(* CODESYS project CanOpen.project
   Title: Opus30
   Version: 1.0.0.0
   Author: Marcus Adolfi
   Company: Schneider Electric

Project tree, tasks and I/O mapping:
  MyController : TM241CE40T/U, Schneider Electric, order no. TM241CE40T/U, version 4.0.2.20
    application Application
      libraries: SysTime, 3.4.1.20 (System)
      task MAST (cyclic, interval 10 ms, priority 15, watchdog 100 ms x 1) calls R00_main
      task VISU_TASK (cyclic, interval 100 ms, priority 30) calls VisuElems.Visu_Prg
      task Task1ms (cyclic, interval 1 ms, priority 1) calls F04_foto, D04_foto, S06_seguranca
      global variables GVL
      01_Machine/
        program R06_principal [LD]
        program R01_firstScan [LD]
        program R05_comando [LD]
        program R21_estatistica [ST]
        program R22_velocMedia [ST]
        program R98_paramFab [ST]
        program R20_acessorios [LD]
        program R99_calcTempos [ST]
        program R00_main [LD]
      Structs/
        data type _exec_bits
        data type _eixo_drive
        data type _eixo_home
        data type _eixo_auto
        data type _receita
        data type _eixo
        data type _bio
        data type _oee
        data type _prev
      05_IHM/
        program I02_alarmes [ST]
        program I07_procedimento [LD]
        program I06_textoConfirma [LD]
        program I01_geral [LD]
        program I03_mensagens [ST]
      02_Filme/
        program F99_calculo [ST]
        program F03_auto [LD]
        program F01_geral [LD]
        program F04_foto [LD]
      global variables PersistentVars
      03_Selagem/
        program S02_home [LD]
        program S99_calculo [ST]
        program S06_seguranca [LD]
        program S01_geral [LD]
        program S03_auto [LD]
      global variables IHM
      Symbol configuration
      04_Disco/
        program D99_calculo [ST]
        program D03_auto [LD]
        program D04_foto [LD]
      function HiddenPOU [ST]
      Visu/
        visualisation Info
        visualisation Main
      10_Relogio/
        function block GetDateAndTime [CFC]
        function block SetDateAndTime [CFC]
        program AjustaDataHora [LD]
      image pool Imagens
      11_FB/
        function block RTO [ST]
      06_bio/
        program B01_controle [ST]
        program B02_data [ST]
      07_dados/
        program D01_data [ST]
        program D02_clean [ST]
        program D03_view [ST]
        program D04_controleView [ST]
      08_manut/
        program U01_controle [ST]
        program U02_soma [ST]
        program U03_reset [ST]
        program U04_view [ST]
        program U00_valoresMax [ST]
    Cartridge_1 : Cartridge, Schneider Electric, version 4.0.2.20
    Cartridge_2 : Cartridge, Schneider Electric, version 4.0.2.20
    IO_Bus : IO bus - TM3, Schneider Electric, version 4.0.2.20
    COM_Bus : COM bus, Schneider Electric, version 4.0.2.20
    Ethernet_1 : Ethernet Network, Schneider Electric, version 4.0.2.20
        settings: IPAddress = [192, 168, 1, 10]; SubnetMask = [255, 255, 255, 0]; WebServer = TRUE; FTP Server = TRUE; SoMachine Protocol = TRUE; Modbus Server = TRUE; NetManage Protocol = TRUE; SNMP protocol = TRUE; WebVisu protocol = TRUE
    Serial_Line_1 : Serial line, Schneider Electric, version 4.0.2.20
      SoMachine_Network_Manager : SoMachine-Network Manager, Schneider Electric, version 4.0.0.2
    Serial_Line_2 : Serial line, Schneider Electric, version 4.0.2.20
      Modbus_Manager : Modbus Manager, Schneider Electric, version 4.0.0.7
    DI : Digital Inputs, Schneider Electric, version 4.0.2.20
        input  i_fotoFilme : BOOL  // IDW0.I0
        input  i_selagFechado : BOOL  // IDW0.I1
        input  i_fotoDisco : BOOL  // IDW0.I2
        input  i_segProduto : BOOL  // IDW0.I3
        input  i_fechamDisco : BOOL  // IDW0.I4
        input  i_selagAberto : BOOL  // IDW0.I5
        input  i_paradaCorte : BOOL  // IDW0.I6
        input  i_relePortaSeg : BOOL  // IDW0.I7
        input  i_segParada : BOOL  // IDW0.I8
        input  i_btReset : BOOL  // IDW0.I9
        input  i_releEmergencia : BOOL  // IDW0.I10
        input  i_marchaAutomatica : BOOL  // IDW0.I11
        input  i_botaoCiclo : BOOL  // IDW0.I12
        input  i_falhaTemperatura : BOOL  // IDW0.I13
        input  i_falhaImpressora : BOOL  // IDW0.I14
        unmapped channels: IDW0, IB1
    DQ : Digital Outputs, Schneider Electric, version 4.0.2.20
        output o_corte : BOOL  // QW0.Q6
        output o_impressao : BOOL  // QW0.Q7
        output o_compressor : BOOL  // QW0.Q9
        output o_injecaoAr : BOOL  // QW0.Q10
        output o_liberaFilme : BOOL  // QW0.Q13
        output qbDQ_QB1 : BYTE  // QB1
        unmapped channels: QW0
    Counters : Counters, Schneider Electric, version 4.0.2.20
    Pulse_Generators : Pulse Generators, Schneider Electric, version 4.0.2.20
        settings: InstanceNumber = 0; Instance name = 'filme_PTO'; Temporary Instance name = 'filme_PTO'; InstanceNumber = 1; Instance name = 'selag_PTO'; Temporary Instance name = 'selag_PTO'
  HMISTU855 : HMIS5T, Schneider Electric, order no. HMIS5T, version 3.5.3.46
    HMI Application
    Ethernet
      SoMachine_Network_Manager2 : SoMachine-Network Manager, Schneider Electric, version 4.0.0.2
    USB
      SoMachine_Network_Manager3 : SoMachine-Network Manager, Schneider Electric, version 4.0.0.2
    COM1
      SoMachine_Network_Manager1 : SoMachine-Network Manager, Schneider Electric, version 4.0.0.2
  6c0f7fb6-600b-4c93-9262-20cdc603757e
  text list GlobalTextList
  5ce3da45-db07-42e7-a21c-a00fff4ed8f6|C:\_Clientes\Opuspac\Doc\Figuras\Botao.png
  5ce3da45-db07-42e7-a21c-a00fff4ed8f6|C:\_Clientes\Opuspac\Doc\Figuras\Botao_ps.png
  5ce3da45-db07-42e7-a21c-a00fff4ed8f6|C:\_Clientes\Opuspac\Doc\Figuras\LogoOpus.jpg
*)

// MyController/Application/Structs/_exec_bits
TYPE _exec_bits :
STRUCT
	RQ					: BOOL;
	IP					: BOOL;
	DN					: BOOL;
	Fase				: DINT;
	Mask				: DINT;
END_STRUCT
END_TYPE

// MyController/Application/Structs/_eixo_drive
TYPE _eixo_drive :
STRUCT
	falha			: MC_ReadAxisError_PTO;
	posicao			: MC_ReadActualPosition_PTO;
	power			: MC_Power_PTO;
	reset			: MC_Reset_PTO;
	status			: MC_ReadMotionState_PTO;
	stop			: MC_Stop_PTO;
END_STRUCT
END_TYPE

// MyController/Application/Structs/_eixo_home
TYPE _eixo_home :
STRUCT
	RQ					: BOOL;
	IP					: BOOL;
	DN					: BOOL;
	Fase				: DINT;
	Mask				: DINT;
	movVeloc			: MC_MoveVelocity_PTO;
	movRelat			: MC_MoveRelative_PTO;
	movStop				: ARRAY[1..2] OF MC_Stop_PTO;
	setPos				: MC_SetPosition_PTO;
END_STRUCT
END_TYPE

// MyController/Application/Structs/_eixo_auto
TYPE _eixo_auto :
STRUCT
	movVeloc					: MC_MoveVelocity_PTO;
	movAbs						: ARRAY[0..2] OF MC_MoveAbsolute_PTO;
	movRelat					: ARRAY[0..2] OF MC_MoveRelative_PTO;
	movStop						: MC_Stop_PTO;
	setPos						: MC_SetPosition_PTO;
END_STRUCT
END_TYPE

// MyController/Application/Structs/_receita
TYPE _receita :
STRUCT
	inicioAtraso				: DINT;

	// Filme
	filmeExtra					: BOOL;
	filmeMmAposFoto				: DINT;
	filmeMmExtra				: DINT;
	
	// Disco
	discoMmAposFoto				: DINT;
	discoAtraso					: DINT;
END_STRUCT
END_TYPE

// MyController/Application/Structs/_eixo
TYPE _eixo :
STRUCT
	auto				: _eixo_auto;
	home				: _eixo_home;
	drive				: _eixo_drive;
	falha				: BOOL;
	posicaoAtual		: DINT;
	calcula				: BOOL;
END_STRUCT
END_TYPE

// MyController/Application/Structs/_bio
TYPE _bio :
STRUCT
	login						: WSTRING:= "";
	loginData					: BOOL;
	bioData						: ARRAY [0..49] OF DINT;
	bioHora						: ARRAY [0..49] OF DINT;
	bioMin						: ARRAY [0..49] OF DINT;
	bioUser						: ARRAY [0..49] OF WSTRING;
	bioGui						: ARRAY [0..49] OF BOOL;
	iz							: DINT:= 0;
END_STRUCT
END_TYPE

// MyController/Application/Structs/_oee
TYPE _oee :
STRUCT
	produtividade				: ARRAY [0..30] OF REAL;
	diaProduzido				: ARRAY [0..30] OF UINT;
	horasProduzidas				: ARRAY [0..30] OF DINT;
	minProduzidos				: ARRAY [0..30] OF DINT;
	diaProduzindo				: DINT;
	mesProduzindo				: DINT;
	anoProduzindo				: DINT;
	backUpdia					: BOOL;
	pontIhm						: ARRAY [0..30] OF BOOL;
	diaProd						: DINT;
END_STRUCT
END_TYPE

// MyController/Application/Structs/_prev
TYPE _prev :
STRUCT
	M_ciclosMax	 				: ARRAY[ 0..7] OF  DINT;
	ciclos						: ARRAY[ 0..7] OF  DINT;
	msg							: ARRAY[ 0..7] OF  BOOL;
	habilita					: ARRAY[ 0..7] OF BOOL;
END_STRUCT
END_TYPE

// MyController/Application/GVL
VAR_GLOBAL
	// transições
	psBtCiclo					: BOOL;

	// Variaveis gerais
	alarmeReset					: BOOL;
	alarmeResetInd				: BOOL;
	alarmeResetBtn				: BOOL;
	alwaysOff					: BOOL;
	alwaysOn					: BOOL;
	arOK						: BOOL;
	biometricoOk				: BOOL;
	calcGeral					: BOOL;
	calcTempos					: BOOL;
	comandoOff					: BOOL;
	contaReset					: BOOL;
	emergOk						: BOOL;
	estatReset					: BOOL;
	existeAlarme				: BOOL;
	falhaImpressora				: BOOL;
	falhaProduto				: BOOL;
	falhaSensorProd				: BOOL;
	falhaTemperatura			: BOOL;
	firstScan					: BOOL;
	injecaoTpoOff				: BOOL;
	liberaCiclo					: BOOL;
	livreComando				: BOOL;
	livreStart					: BOOL;
	modoAutomatico				: BOOL;					
	pisca						: BOOL;
	piscaRapido					: BOOL;
	primeiroCiclo				: BOOL;
	setAmpola					: BOOL;
	tpoDisco					: TIME;
	tpoInicio					: TIME;
	tpoInjecao					: TIME;
	tpoSelagem					: TIME;
	
	
	
	TL_inicializa				: TON;
	TL_disco					: TON;
	TF_corte					: TON;
	
	acopla						: _exec_bits;
	ciclo						: _exec_bits;
	comando						: _exec_bits;
	compressor					: _exec_bits;
	conta						: _exec_bits;
	corte						: _exec_bits;
	injecaoAr					: _exec_bits;
	media						: _exec_bits;
	mudaReceita					: _exec_bits;
	principal					: _exec_bits;
	vidaUtil					: _exec_bits;
	
	// Alimentador de Blisters
	msgPrimeiro					: BOOL;
	limpaDados					: BOOL;
	procedimento				: ARRAY[0..2] OF _exec_bits;

	
	// Variaveis Filme
	filme						: _eixo;
	filmeMove					: ARRAY[0..2] OF _exec_bits;
	filmeParaImed				: BOOL;
	filmeVeloc					: DINT;
	filmeExtra					: BOOL;
	filmeFotoOk					: BOOL;
	filmePulsosAposFoto			: DINT;
	filmePulsosExtra			: DINT;
	filmePulsosMm				: REAL;
	filmePreso					: _exec_bits;
	
	// Variaveis Selagem
	selag						: _eixo;
	selagAbre					: _exec_bits;
	selagFecha					: _exec_bits;
	selagVeloc					: DINT;
	selagVelocHome				: DINT;
	selagPulsosMm				: REAL;
	selagPulsosFechar			: DINT;

	// Variaveis Disco
	disco						: _eixo;
	discoMove					: _exec_bits;
	discoParaImed				: BOOL;
	discoVeloc					: DINT;
	discoPulsosMm				: REAL;
	discoPulsosAposFoto			: DINT;
	
	// Variaveis Visualization
	vsBtStart					: BOOL;
	vsMarchaAutomatica			: BOOL;
	
	
    //Sincroniza e ajusta o relógio da IHM
	AnoSet						: UINT;
	ClkScan						: BOOL;
	AjustaHora					: BOOL;
	MesSet						: UINT;
	DiaSet						: UINT;
	HoraSet						: UINT;
	MinutoSet					: UINT;
	SegundoSet					: UINT;
	AnoAtual					: UINT;
	MesAtual					: UINT;
	DiaAtual					: UINT;
	HoraAtual					: UINT;
	MinutoAtual					: UINT;
	SegundoAtual				: UINT;	
	sink						: BOOL;

	
(*	=================== ALARMES ===================
	Obs: alarme[0]- Não utilizado
*)
	alarme						: ARRAY[0..50] OF BOOL;
	alarmes						: _exec_bits;
	mensagem					: ARRAY[0..50] OF BOOL;
	numAlarme					: SINT;
END_VAR

// MyController/Application/PersistentVars
VAR_GLOBAL PERSISTENT RETAIN
	versaoSoftware				: REAL:= 1.00;
	pi							: REAL:= 3.1415926;
	paramFab					: BOOL:= TRUE;
	contaAtual					: DINT;
	contaGeral					: DINT;
	contaSet					: DINT;
	numReceita					: SINT;
	
	M_tpoInjecaoAr				: DINT:= 99;
	M_produtMedio				: DINT:= 70;
	M_tpoFormato				: TIME:= T#280MS;
	
	// Informações
	infoTpoEnergHrs				: DINT;
	infoTpoEnergMin				: DINT;
	infoTpoProdHrs				: DINT;
	infoTpoProdMin				: DINT;
	
	// Filme
	M_filmePulsosVolta			: DINT:= 1600;
	M_diamRolo					: DINT:= 34;
	M_filmeVeloc				: DINT:= 40;
	M_filmeAcel					: DINT:= 200;
	M_filmeDecel				: DINT:= 100;
	
	// Disco
	M_discoPulsosVolta			: DINT:= 6400;
	M_diamDisco					: DINT:= 166;
	M_discoVeloc				: DINT:= 4;
	M_discoAcel					: DINT:= 150;
	M_discoDecel				: DINT:= 150;
	
	// Selagem
	M_selagPulsosVolta			: DINT:= 20000;
	M_selagVelocHome			: DINT:= 20;
	M_selagVeloc				: DINT:= 100;
	M_selagTpoSelagem			: DINT:= 20;
	M_selagPosFecha				: DINT:= 789;
	M_selagAcel					: DINT:= 40;
	M_selagDecel				: DINT:= 40;
	
	// Receita
	Rc							: ARRAY[0..3] OF _receita;
	Fb							: ARRAY[0..3] OF _receita;
	
	// IHM
	ihm_procedCurto				: BOOL;
	
	// Digital
	digital						: _bio;
	iz							: DINT;
	
	// biometria
	ihm_digitalInstalado		: BOOL;
	
	// Dados
	dados						: _oee;
	indPainel					: DINT:= 0;
	indSub						: BOOL;
	indSoma						: BOOL;
	panData						: ARRAY [0..08] OF DINT;
	panProd						: ARRAY [0..08] OF REAL;
	panHora						: ARRAY [0..08] OF DINT;
	panMin						: ARRAY [0..08] OF DINT;
	pt							: DINT:= 0;
	pa							: DINT;
	
	// Vida Util
	util						: _prev; 
END_VAR

// MyController/Application/IHM
VAR_GLOBAL
	ihm_alarme					: ARRAY[0..50] OF BOOL;
	ihm_alarmeReset				: BOOL;
	ihm_alarmeResetInd			: BOOL;
	ihm_bannerConfirma			: BOOL;
	ihm_bannerMensagem			: BOOL;
	ihm_carregaFabrica			: BOOL;
	ihm_confirmaV				: BOOL;
	ihm_confirmaX				: BOOL;
	ihm_contaAtual				: DINT;
	ihm_contaGeral				: DINT;
	ihm_contaReset				: BOOL;
	ihm_entrada					: ARRAY[0..23] OF BOOL;
	ihm_estatReset				: BOOL;
	ihm_mensagem				: DINT;
	ihm_numReceita				: SINT;
	ihm_preso					: BOOL;
	ihm_produtMedio				: REAL;
	ihm_telaHome				: BOOL;
	ihm_salvaFabrica			: BOOL;
	ihm_saida					: ARRAY[0..15] OF BOOL;
	ihm_selagHome				: BOOL;
	ihm_telaAtual				: INT;
	ihm_textoConfirma			: DINT;
	ihm_textoProced				: DINT;
	ihm_velocMedida				: DINT;
	ihm_visibPhone				: BOOL;
	ihm_setUpAmpola				: BOOL;
	
	// Produtividade
	ihm_backUpProdutividade		: BOOL;
	
	
	ihm_digitalHabilitado		: BOOL;
	ihm_usuarioLoggado			: BOOL;
	ihm_realizaBackup 			: BOOL;	
	
	// Vida Util 
	ihm_resetCiclos				: ARRAY[0..7] OF BOOL;
END_VAR

// MyController/Application/01_Machine/R00_main
PROGRAM R00_main
VAR
END_VAR

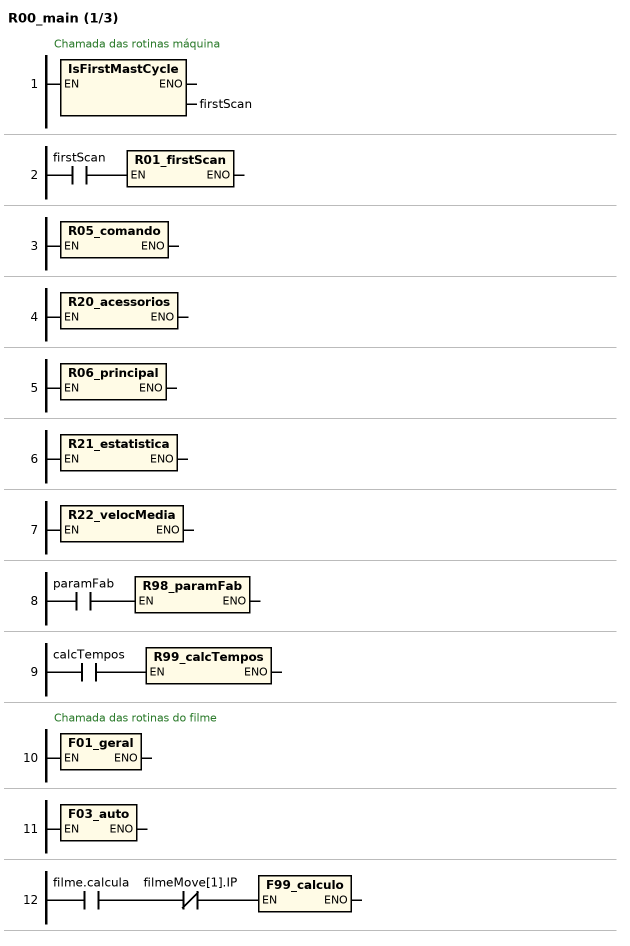
// NETWORK 1
// Chamada das rotinas máquina
firstScan := IsFirstMastCycle();

// NETWORK 2
IF firstScan THEN R01_firstScan(); END_IF

// NETWORK 3
R05_comando();

// NETWORK 4
R20_acessorios();

// NETWORK 5
R06_principal();

// NETWORK 6
R21_estatistica();

// NETWORK 7
R22_velocMedia();

// NETWORK 8
IF paramFab THEN R98_paramFab(); END_IF

// NETWORK 9
IF calcTempos THEN R99_calcTempos(); END_IF

// NETWORK 10
// Chamada das rotinas do filme
F01_geral();

// NETWORK 11
F03_auto();

// NETWORK 12
IF filme.calcula AND NOT filmeMove[1].IP THEN F99_calculo(); END_IF

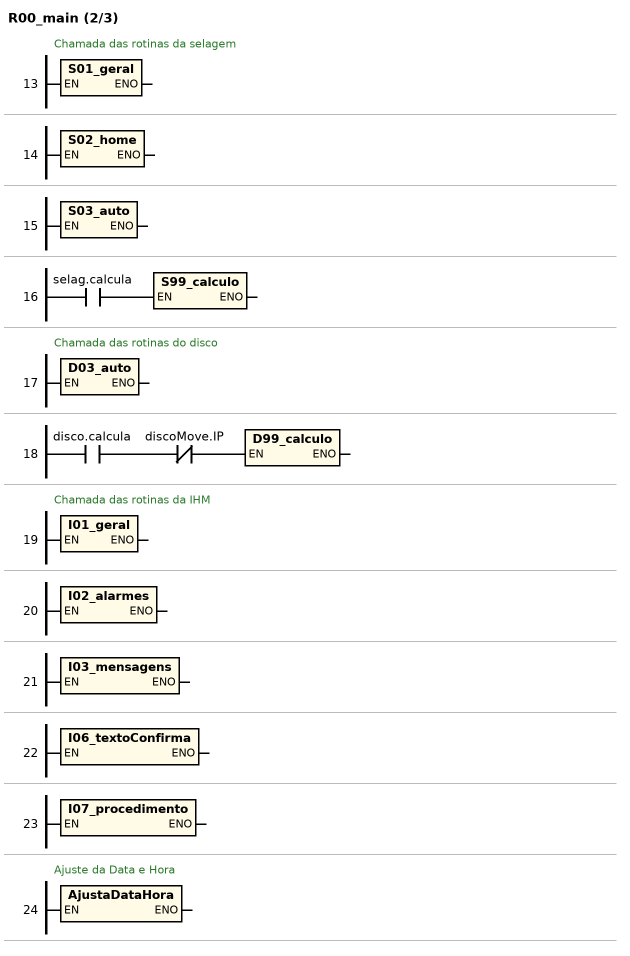
// NETWORK 13
// Chamada das rotinas da selagem
S01_geral();

// NETWORK 14
S02_home();

// NETWORK 15
S03_auto();

// NETWORK 16
IF selag.calcula THEN S99_calculo(); END_IF

// NETWORK 17
// Chamada das rotinas do disco
D03_auto();

// NETWORK 18
IF disco.calcula AND NOT discoMove.IP THEN D99_calculo(); END_IF

// NETWORK 19
// Chamada das rotinas da IHM
I01_geral();

// NETWORK 20
I02_alarmes();

// NETWORK 21
I03_mensagens();

// NETWORK 22
I06_textoConfirma();

// NETWORK 23
I07_procedimento();

// NETWORK 24
// Ajuste da Data e Hora
AjustaDataHora();

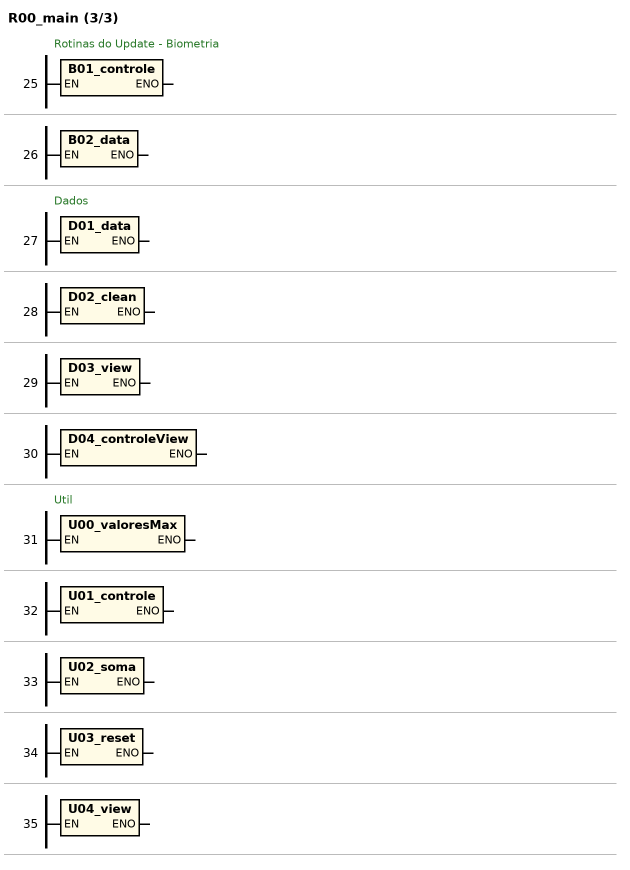
// NETWORK 25
// Rotinas do Update - Biometria
B01_controle();

// NETWORK 26
B02_data();

// NETWORK 27
//     Dados
D01_data();

// NETWORK 28
D02_clean();

// NETWORK 29
D03_view();

// NETWORK 30
D04_controleView();

// NETWORK 31
// Util
U00_valoresMax();

// NETWORK 32
U01_controle();

// NETWORK 33
U02_soma();

// NETWORK 34
U03_reset();

// NETWORK 35
U04_view();

END_PROGRAM

// MyController/Application/01_Machine/R01_firstScan
PROGRAM R01_firstScan
VAR
END_VAR

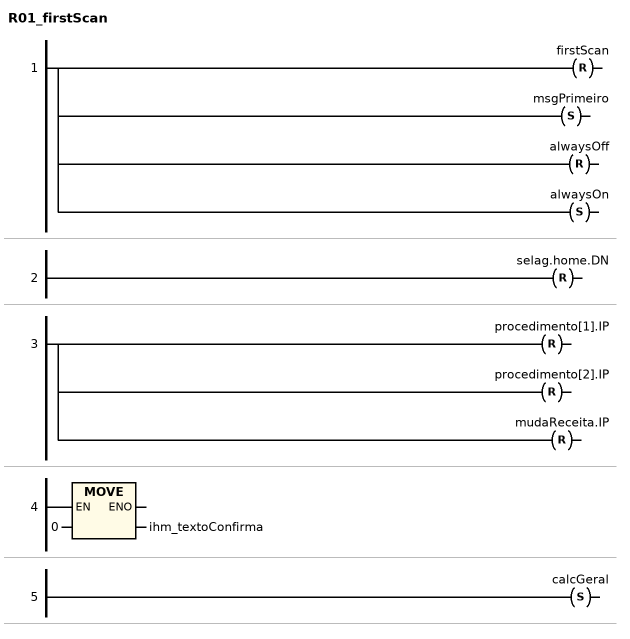
// NETWORK 1
firstScan R= TRUE;
msgPrimeiro S= TRUE;
alwaysOff R= TRUE;
alwaysOn S= TRUE;

// NETWORK 2
selag.home.DN R= TRUE;

// NETWORK 3
procedimento[1].IP R= TRUE;
procedimento[2].IP R= TRUE;
mudaReceita.IP R= TRUE;

// NETWORK 4
ihm_textoConfirma := 0;

// NETWORK 5
calcGeral S= TRUE;

END_PROGRAM

// MyController/Application/01_Machine/R05_comando
PROGRAM R05_comando
VAR
	TL_comando				: TON;
END_VAR
VAR // added by the converter: edge detectors and wires of the graphical bodies
    _rt1, _rt2, _rt3, _rt4 : R_TRIG;
    _w1, _w2 : BOOL;
    _ft1, _ft2, _ft3 : F_TRIG;
END_VAR

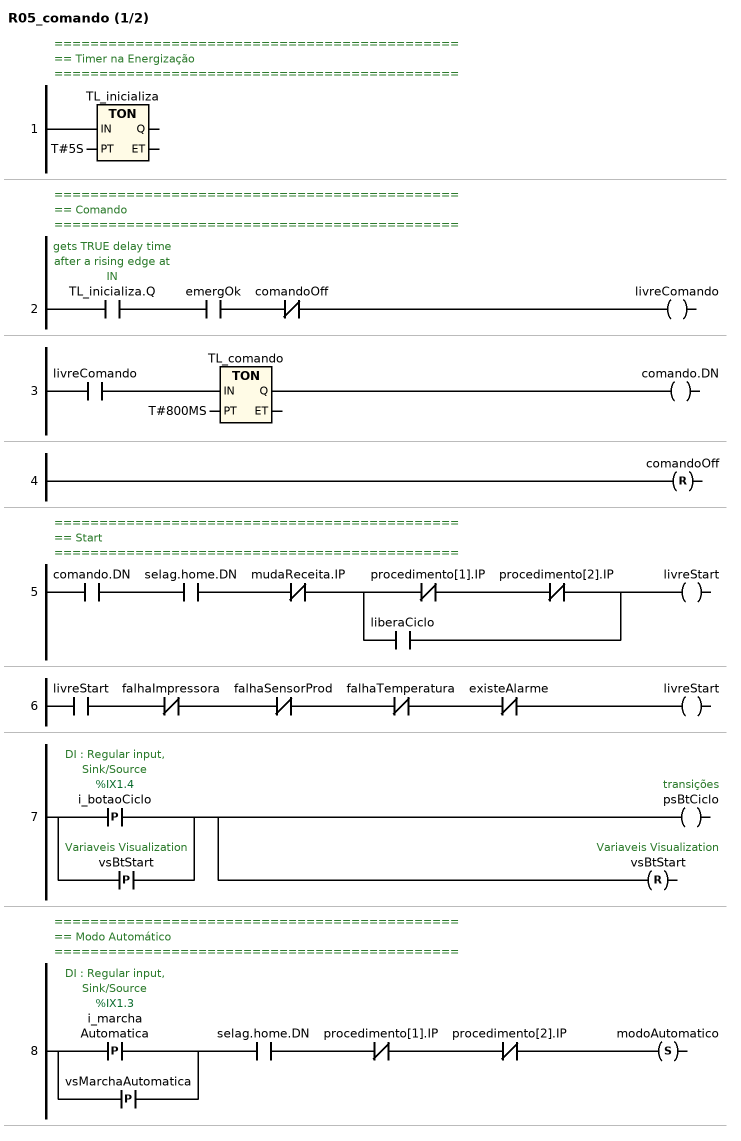
// NETWORK 1
// =============================================
// == Timer na Energização
// =============================================
TL_inicializa(IN := TRUE, PT := T#5S); // TON

// NETWORK 2
// =============================================
// == Comando
// =============================================
//   TL_inicializa.Q: gets TRUE delay time after a rising edge at IN
livreComando := TL_inicializa.Q AND emergOk AND NOT comandoOff;

// NETWORK 3
TL_comando(IN := livreComando, PT := T#800MS); // TON
comando.DN := TL_comando.Q;

// NETWORK 4
comandoOff R= TRUE;

// NETWORK 5
// =============================================
// == Start
// =============================================
livreStart := comando.DN AND selag.home.DN AND NOT mudaReceita.IP AND (NOT procedimento[1].IP AND NOT procedimento[2].IP OR liberaCiclo);

// NETWORK 6
livreStart := livreStart AND NOT falhaImpressora AND NOT falhaSensorProd AND NOT falhaTemperatura AND NOT existeAlarme;

// NETWORK 7
//   i_botaoCiclo: DI : Regular input, Sink/Source | AT %IX1.4
//   vsBtStart: Variaveis Visualization
//   psBtCiclo: transições
_rt1(CLK := i_botaoCiclo);
_rt2(CLK := vsBtStart);
_w1 := _rt1.Q OR _rt2.Q;
psBtCiclo := _w1;
vsBtStart R= _w1;

// NETWORK 8
// =============================================
// == Modo Automático
// =============================================
//   i_marchaAutomatica: DI : Regular input, Sink/Source | AT %IX1.3
_rt3(CLK := i_marchaAutomatica);
_rt4(CLK := vsMarchaAutomatica);
modoAutomatico S= (_rt3.Q OR _rt4.Q) AND selag.home.DN AND NOT procedimento[1].IP AND NOT procedimento[2].IP;

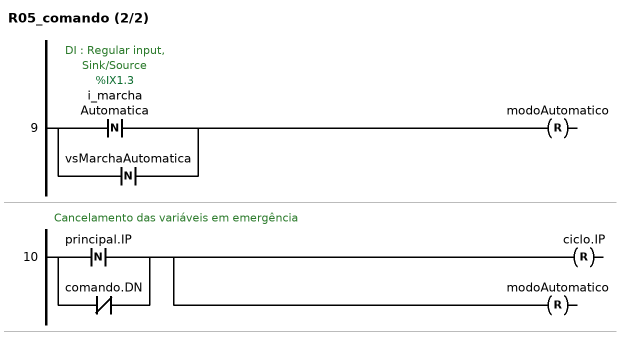
// NETWORK 9
//   i_marchaAutomatica: DI : Regular input, Sink/Source | AT %IX1.3
_ft1(CLK := i_marchaAutomatica);
_ft2(CLK := vsMarchaAutomatica);
modoAutomatico R= _ft1.Q OR _ft2.Q;

// NETWORK 10
// Cancelamento das variáveis em emergência
_ft3(CLK := principal.IP);
_w2 := _ft3.Q OR NOT comando.DN;
ciclo.IP R= _w2;
modoAutomatico R= _w2;

END_PROGRAM

// MyController/Application/01_Machine/R20_acessorios
PROGRAM R20_acessorios
VAR
	TD_injecaoAr				: TON;
	TD_compressor				: TON;
	TL_compressor				: TON;
	TL_filmePreso				: TON;
	TF_impressora				: TON;
	TL_pisca					: BLINK;
	TL_piscaRapido				: BLINK;
	TF_temperatura				: TON;
END_VAR
VAR // added by the converter: edge detectors and wires of the graphical bodies
    _w1, _w2, _w3, _w4 : BOOL;
    _rt1, _rt2, _rt3 : R_TRIG;
    _ft1, _ft2, _ft3 : F_TRIG;
END_VAR

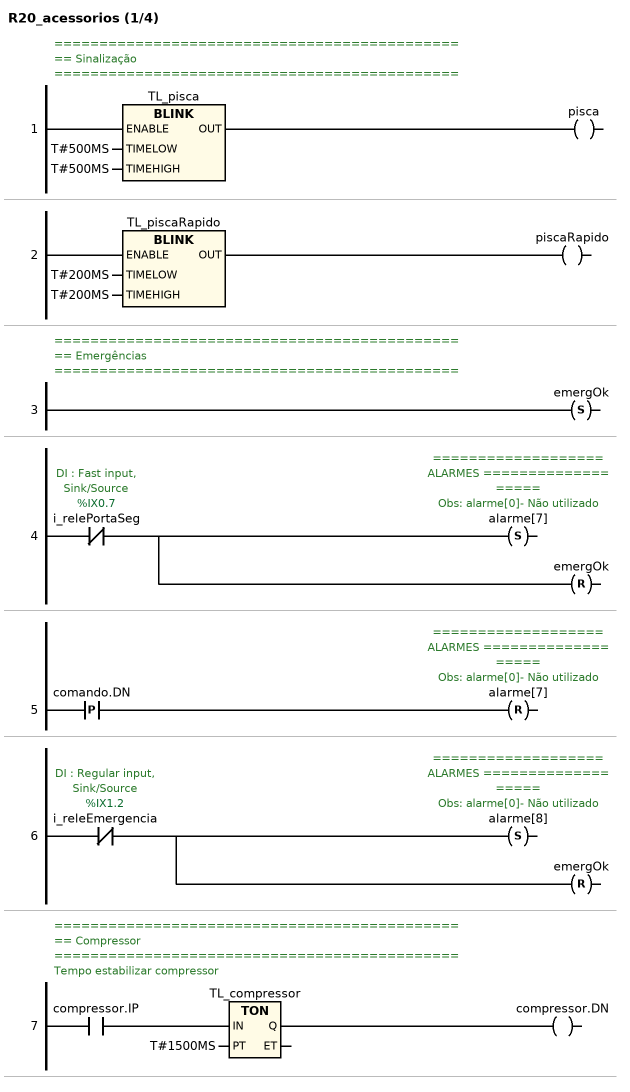
// NETWORK 1
// =============================================
// == Sinalização
// =============================================
TL_pisca(ENABLE := TRUE, TIMELOW := T#500MS, TIMEHIGH := T#500MS); // BLINK
pisca := TL_pisca.OUT;

// NETWORK 2
TL_piscaRapido(ENABLE := TRUE, TIMELOW := T#200MS, TIMEHIGH := T#200MS); // BLINK
piscaRapido := TL_piscaRapido.OUT;

// NETWORK 3
// =============================================
// == Emergências
// =============================================
emergOk S= TRUE;

// NETWORK 4
//   i_relePortaSeg: DI : Fast input, Sink/Source | AT %IX0.7
//   alarme[7]: =================== ALARMES =================== Obs: alarme[0]- Não utilizado
_w1 := NOT i_relePortaSeg;
alarme[7] S= _w1;
emergOk R= _w1;

// NETWORK 5
//   alarme[7]: =================== ALARMES =================== Obs: alarme[0]- Não utilizado
_rt1(CLK := comando.DN);
alarme[7] R= _rt1.Q;

// NETWORK 6
//   i_releEmergencia: DI : Regular input, Sink/Source | AT %IX1.2
//   alarme[8]: =================== ALARMES =================== Obs: alarme[0]- Não utilizado
_w2 := NOT i_releEmergencia;
alarme[8] S= _w2;
emergOk R= _w2;

// NETWORK 7
// =============================================
// == Compressor
// =============================================
// Tempo estabilizar compressor
TL_compressor(IN := compressor.IP, PT := T#1500MS); // TON
compressor.DN := TL_compressor.Q;

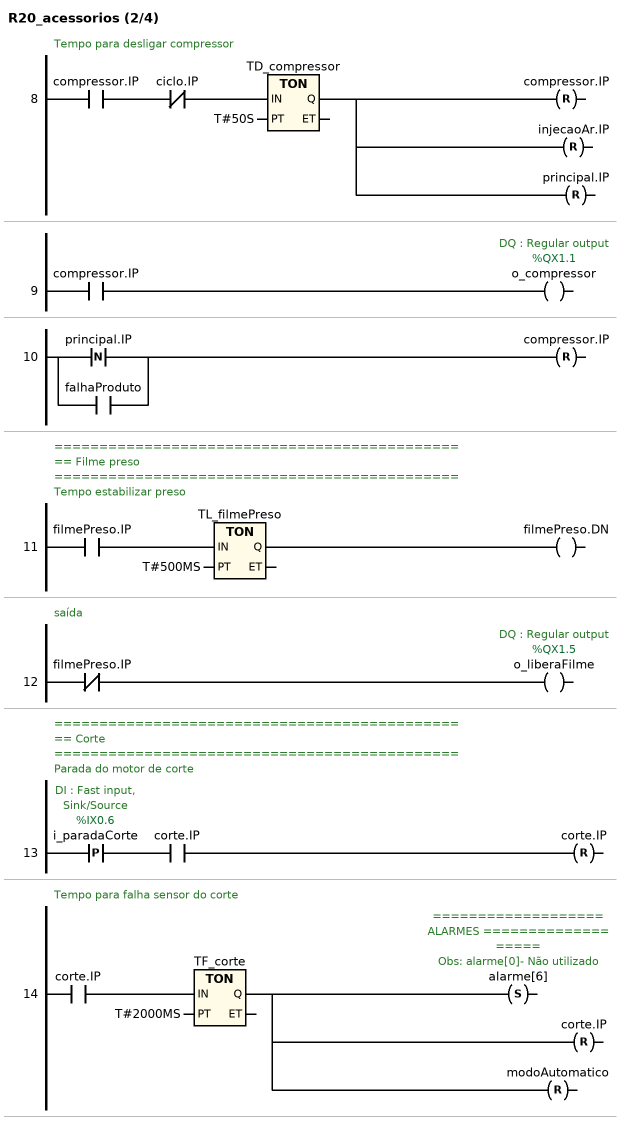
// NETWORK 8
// Tempo para desligar compressor
TD_compressor(IN := compressor.IP AND NOT ciclo.IP, PT := T#50S); // TON
compressor.IP R= TD_compressor.Q;
injecaoAr.IP R= TD_compressor.Q;
principal.IP R= TD_compressor.Q;

// NETWORK 9
//   o_compressor: DQ : Regular output | AT %QX1.1
o_compressor := compressor.IP;

// NETWORK 10
_ft1(CLK := principal.IP);
compressor.IP R= _ft1.Q OR falhaProduto;

// NETWORK 11
// =============================================
// == Filme preso
// =============================================
// Tempo estabilizar preso
TL_filmePreso(IN := filmePreso.IP, PT := T#500MS); // TON
filmePreso.DN := TL_filmePreso.Q;

// NETWORK 12
// saída
//   o_liberaFilme: DQ : Regular output | AT %QX1.5
o_liberaFilme := NOT filmePreso.IP;

// NETWORK 13
// =============================================
// == Corte
// =============================================
// Parada do motor de corte
//   i_paradaCorte: DI : Fast input, Sink/Source | AT %IX0.6
_rt2(CLK := i_paradaCorte);
corte.IP R= _rt2.Q AND corte.IP;

// NETWORK 14
// Tempo para falha sensor do corte
//   alarme[6]: =================== ALARMES =================== Obs: alarme[0]- Não utilizado
TF_corte(IN := corte.IP, PT := T#2000MS); // TON
alarme[6] S= TF_corte.Q;
corte.IP R= TF_corte.Q;
modoAutomatico R= TF_corte.Q;

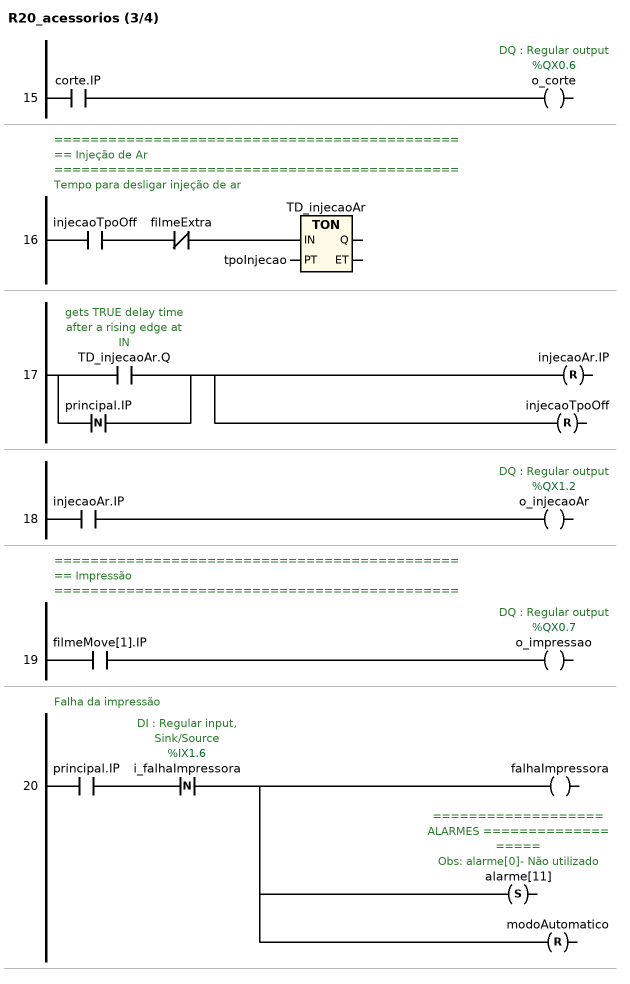
// NETWORK 15
//   o_corte: DQ : Regular output | AT %QX0.6
o_corte := corte.IP;

// NETWORK 16
// =============================================
// == Injeção de Ar
// =============================================
// Tempo para desligar injeção de ar
TD_injecaoAr(IN := injecaoTpoOff AND NOT filmeExtra, PT := tpoInjecao); // TON

// NETWORK 17
//   TD_injecaoAr.Q: gets TRUE delay time after a rising edge at IN
_ft2(CLK := principal.IP);
_w3 := TD_injecaoAr.Q OR _ft2.Q;
injecaoAr.IP R= _w3;
injecaoTpoOff R= _w3;

// NETWORK 18
//   o_injecaoAr: DQ : Regular output | AT %QX1.2
o_injecaoAr := injecaoAr.IP;

// NETWORK 19
// =============================================
// == Impressão
// =============================================
//   o_impressao: DQ : Regular output | AT %QX0.7
o_impressao := filmeMove[1].IP;

// NETWORK 20
// Falha da impressão
//   i_falhaImpressora: DI : Regular input, Sink/Source | AT %IX1.6
//   alarme[11]: =================== ALARMES =================== Obs: alarme[0]- Não utilizado
_ft3(CLK := i_falhaImpressora);
_w4 := principal.IP AND _ft3.Q;
falhaImpressora := _w4;
alarme[11] S= _w4;
modoAutomatico R= _w4;

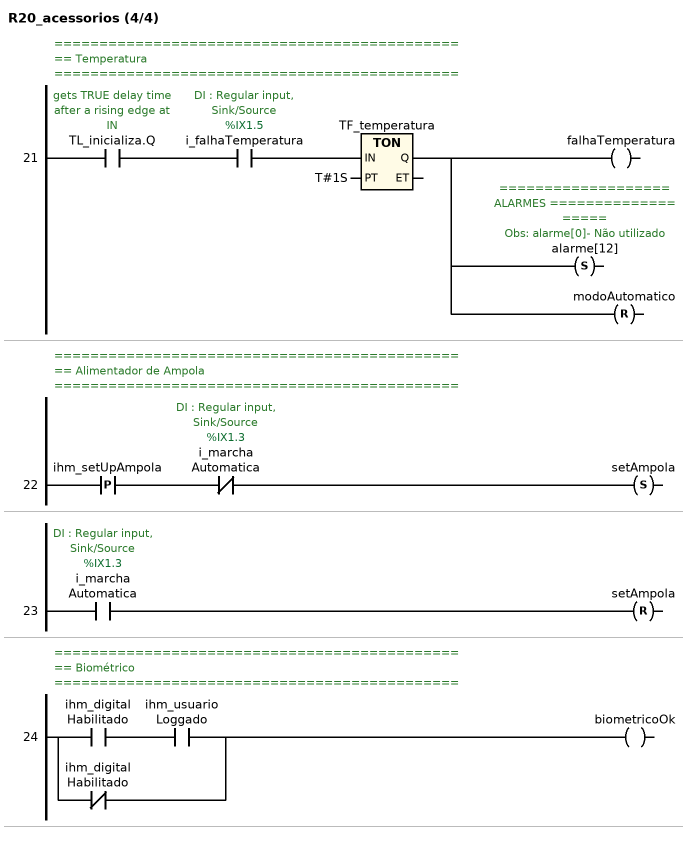
// NETWORK 21
// =============================================
// == Temperatura
// =============================================
//   TL_inicializa.Q: gets TRUE delay time after a rising edge at IN
//   i_falhaTemperatura: DI : Regular input, Sink/Source | AT %IX1.5
//   alarme[12]: =================== ALARMES =================== Obs: alarme[0]- Não utilizado
TF_temperatura(IN := TL_inicializa.Q AND i_falhaTemperatura, PT := T#1S); // TON
falhaTemperatura := TF_temperatura.Q;
alarme[12] S= TF_temperatura.Q;
modoAutomatico R= TF_temperatura.Q;

// NETWORK 22
// =============================================
// == Alimentador de Ampola
// =============================================
//   i_marchaAutomatica: DI : Regular input, Sink/Source | AT %IX1.3
_rt3(CLK := ihm_setUpAmpola);
setAmpola S= _rt3.Q AND NOT i_marchaAutomatica;

// NETWORK 23
//   i_marchaAutomatica: DI : Regular input, Sink/Source | AT %IX1.3
setAmpola R= i_marchaAutomatica;

// NETWORK 24
// =============================================
// == Biométrico
// =============================================
biometricoOk := ihm_digitalHabilitado AND ihm_usuarioLoggado OR NOT ihm_digitalHabilitado;

END_PROGRAM

// MyController/Application/01_Machine/R06_principal
PROGRAM R06_principal
VAR
	primeiroCiclo			: BOOL;
	execMedida				: _exec_bits;
	tpoMedido				: TIME;
	T_medidaForm			: TON;
	T_inicio				: ARRAY[1..2] OF TON;
	T_selagem				: TON;
	
	T_teste					: TON;
END_VAR
VAR // added by the converter: edge detectors and wires of the graphical bodies
    _w1, _w2, _w3, _w4, _w5, _w6, _w7, _w8, _w9, _w10, _w11, _w12, _w13, _w14, _w15, _w16, _w17, _w18, _w19, _w20, _w21, _w22, _w23 : BOOL;
    _ft1, _ft2 : F_TRIG;
END_VAR

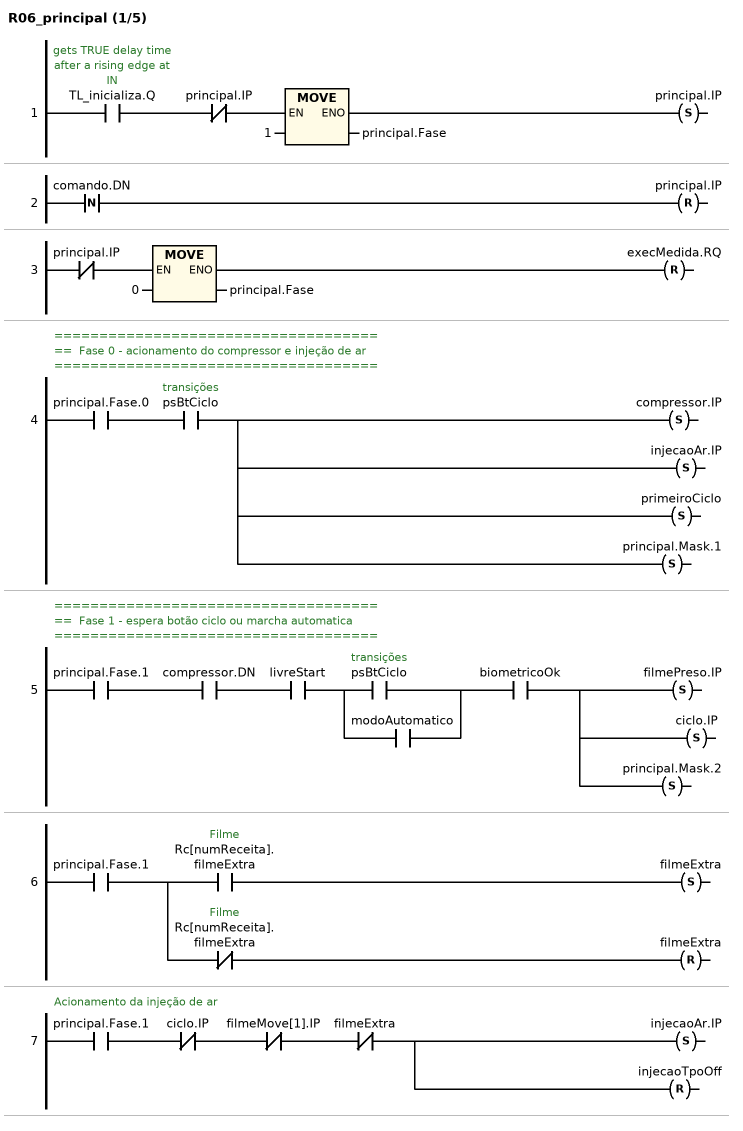
// NETWORK 1
//   TL_inicializa.Q: gets TRUE delay time after a rising edge at IN
_w1 := TL_inicializa.Q AND NOT principal.IP;
IF _w1 THEN principal.Fase := 1; END_IF
principal.IP S= _w1;

// NETWORK 2
_ft1(CLK := comando.DN);
principal.IP R= _ft1.Q;

// NETWORK 3
_w2 := NOT principal.IP;
IF _w2 THEN principal.Fase := 0; END_IF
execMedida.RQ R= _w2;

// NETWORK 4
// ====================================
// ==  Fase 0 - acionamento do compressor e injeção de ar
// ====================================
//   psBtCiclo: transições
_w3 := principal.Fase.0 AND psBtCiclo;
compressor.IP S= _w3;
injecaoAr.IP S= _w3;
primeiroCiclo S= _w3;
principal.Mask.1 S= _w3;

// NETWORK 5
// ====================================
// ==  Fase 1 - espera botão ciclo ou marcha automatica
// ====================================
//   psBtCiclo: transições
_w4 := principal.Fase.1 AND compressor.DN AND livreStart AND (psBtCiclo OR modoAutomatico) AND biometricoOk;
filmePreso.IP S= _w4;
ciclo.IP S= _w4;
principal.Mask.2 S= _w4;

// NETWORK 6
//   Rc[numReceita].filmeExtra: Filme
filmeExtra S= principal.Fase.1 AND Rc[numReceita].filmeExtra;
filmeExtra R= principal.Fase.1 AND NOT Rc[numReceita].filmeExtra;

// NETWORK 7
// Acionamento da injeção de ar
_w5 := principal.Fase.1 AND NOT ciclo.IP AND NOT filmeMove[1].IP AND NOT filmeExtra;
injecaoAr.IP S= _w5;
injecaoTpoOff R= _w5;
